// TIA Portal project "ETI C 25" (V15.1) (continued)
   PLC_TO_PC.DATA[324] := ' ';
   PLC_TO_PC.DATA[325] := ' ';
   PLC_TO_PC.DATA[326] := ' ';
   PLC_TO_PC.DATA[327] := ' ';
   PLC_TO_PC.DATA[328] := ' ';
   PLC_TO_PC.DATA[329] := ' ';
   PLC_TO_PC.DATA[330] := ' ';
   PLC_TO_PC.DATA[331] := ' ';
   PLC_TO_PC.DATA[332] := ' ';
   PLC_TO_PC.DATA[333] := ' ';
   PLC_TO_PC.DATA[334] := ' ';
   PLC_TO_PC.DATA[335] := ' ';
   PLC_TO_PC.DATA[336] := ' ';
   PLC_TO_PC.DATA[337] := ' ';
   PLC_TO_PC.DATA[338] := ' ';
   PLC_TO_PC.DATA[339] := ' ';
   PLC_TO_PC.DATA[340] := ' ';
   PLC_TO_PC.DATA[341] := ' ';
   PLC_TO_PC.DATA[342] := ' ';
   PLC_TO_PC.DATA[343] := ' ';
   PLC_TO_PC.DATA[344] := ' ';
   PLC_TO_PC.DATA[345] := ' ';
   PLC_TO_PC.DATA[346] := ' ';
   PLC_TO_PC.DATA[347] := ' ';
   PLC_TO_PC.DATA[348] := ' ';
   PLC_TO_PC.DATA[349] := ' ';
   PLC_TO_PC.DATA[350] := ' ';
   PLC_TO_PC.DATA[351] := ' ';
   PLC_TO_PC.DATA[352] := ' ';
   PLC_TO_PC.DATA[353] := ' ';
   PLC_TO_PC.DATA[354] := ' ';
   PLC_TO_PC.DATA[355] := ' ';
   PLC_TO_PC.DATA[356] := ' ';
   PLC_TO_PC.DATA[357] := ' ';
   PLC_TO_PC.DATA[358] := ' ';
   PLC_TO_PC.DATA[359] := ' ';
   PLC_TO_PC.DATA[360] := ' ';
   PLC_TO_PC.DATA[361] := ' ';
   PLC_TO_PC.DATA[362] := ' ';
   PLC_TO_PC.DATA[363] := ' ';
   PLC_TO_PC.DATA[364] := ' ';
   PLC_TO_PC.DATA[365] := ' ';
   PLC_TO_PC.DATA[366] := ' ';
   PLC_TO_PC.DATA[367] := ' ';
   PLC_TO_PC.DATA[368] := ' ';
   PLC_TO_PC.DATA[369] := ' ';
   PLC_TO_PC.DATA[370] := ' ';
   PLC_TO_PC.DATA[371] := ' ';
   PLC_TO_PC.DATA[372] := ' ';
   PLC_TO_PC.DATA[373] := ' ';
   PLC_TO_PC.DATA[374] := ' ';
   PLC_TO_PC.DATA[375] := ' ';
   PLC_TO_PC.DATA[376] := ' ';
   PLC_TO_PC.DATA[377] := ' ';
   PLC_TO_PC.DATA[378] := ' ';
   PLC_TO_PC.DATA[379] := ' ';
   PLC_TO_PC.DATA[380] := ' ';
   PLC_TO_PC.DATA[381] := ' ';
   PLC_TO_PC.DATA[382] := ' ';
   PLC_TO_PC.DATA[383] := ' ';
   PLC_TO_PC.DATA[384] := ' ';
   PLC_TO_PC.DATA[385] := ' ';
   PLC_TO_PC.DATA[386] := ' ';
   PLC_TO_PC.DATA[387] := ' ';
   PLC_TO_PC.DATA[388] := ' ';
   PLC_TO_PC.DATA[389] := ' ';
   PLC_TO_PC.DATA[390] := ' ';
   PLC_TO_PC.DATA[391] := ' ';
   PLC_TO_PC.DATA[392] := ' ';
   PLC_TO_PC.DATA[393] := ' ';
   PLC_TO_PC.DATA[394] := ' ';
   PLC_TO_PC.DATA[395] := ' ';
   PLC_TO_PC.DATA[396] := ' ';
   PLC_TO_PC.DATA[397] := ' ';
   PLC_TO_PC.DATA[398] := ' ';
   PLC_TO_PC.DATA[399] := ' ';
   PLC_TO_PC.DATA[400] := ' ';
   PLC_TO_PC.DATA[401] := ' ';
   PLC_TO_PC.DATA[402] := ' ';
   PLC_TO_PC.DATA[403] := ' ';
   PLC_TO_PC.DATA[404] := ' ';
   PLC_TO_PC.DATA[405] := ' ';
   PLC_TO_PC.DATA[406] := ' ';
   PLC_TO_PC.DATA[407] := ' ';
   PLC_TO_PC.DATA[408] := ' ';
   PLC_TO_PC.DATA[409] := ' ';
   PLC_TO_PC.DATA[410] := ' ';
   PLC_TO_PC.DATA[411] := ' ';
   PLC_TO_PC.DATA[412] := ' ';
   PLC_TO_PC.DATA[413] := ' ';
   PLC_TO_PC.DATA[414] := ' ';
   PLC_TO_PC.DATA[415] := ' ';
   PLC_TO_PC.DATA[416] := ' ';
   PLC_TO_PC.DATA[417] := ' ';
   PLC_TO_PC.DATA[418] := ' ';
   PLC_TO_PC.DATA[419] := ' ';
   PLC_TO_PC.DATA[420] := ' ';
   PLC_TO_PC.DATA[421] := ' ';
   PLC_TO_PC.DATA[422] := ' ';
   PLC_TO_PC.DATA[423] := ' ';
   PLC_TO_PC.DATA[424] := ' ';
   PLC_TO_PC.DATA[425] := ' ';
   PLC_TO_PC.DATA[426] := ' ';
   PLC_TO_PC.DATA[427] := ' ';
   PLC_TO_PC.DATA[428] := ' ';
   PLC_TO_PC.DATA[429] := ' ';
   PLC_TO_PC.DATA[430] := ' ';
   PLC_TO_PC.DATA[431] := ' ';
   PLC_TO_PC.DATA[432] := ' ';
   PLC_TO_PC.DATA[433] := ' ';
   PLC_TO_PC.DATA[434] := ' ';
   PLC_TO_PC.DATA[435] := ' ';
   PLC_TO_PC.DATA[436] := ' ';
   PLC_TO_PC.DATA[437] := ' ';
   PLC_TO_PC.DATA[438] := ' ';
   PLC_TO_PC.DATA[439] := ' ';
   PLC_TO_PC.DATA[440] := ' ';
   PLC_TO_PC.DATA[441] := ' ';
   PLC_TO_PC.DATA[442] := ' ';
   PLC_TO_PC.DATA[443] := ' ';
   PLC_TO_PC.DATA[444] := ' ';
   PLC_TO_PC.DATA[445] := ' ';
   PLC_TO_PC.DATA[446] := ' ';
   PLC_TO_PC.DATA[447] := ' ';
   PLC_TO_PC.DATA[448] := ' ';
   PLC_TO_PC.DATA[449] := ' ';
   PLC_TO_PC.DATA[450] := ' ';
   PLC_TO_PC.DATA[451] := ' ';
   PLC_TO_PC.DATA[452] := ' ';
   PLC_TO_PC.DATA[453] := ' ';
   PLC_TO_PC.DATA[454] := ' ';
   PLC_TO_PC.DATA[455] := ' ';
   PLC_TO_PC.DATA[456] := ' ';
   PLC_TO_PC.DATA[457] := ' ';
   PLC_TO_PC.DATA[458] := ' ';
   PLC_TO_PC.DATA[459] := ' ';
   PLC_TO_PC.DATA[460] := ' ';
   PLC_TO_PC.DATA[461] := ' ';
   PLC_TO_PC.DATA[462] := ' ';
   PLC_TO_PC.DATA[463] := ' ';
   PLC_TO_PC.DATA[464] := ' ';
   PLC_TO_PC.DATA[465] := ' ';
   PLC_TO_PC.DATA[466] := ' ';
   PLC_TO_PC.DATA[467] := ' ';
   PLC_TO_PC.DATA[468] := ' ';
   PLC_TO_PC.DATA[469] := ' ';
   PLC_TO_PC.DATA[470] := ' ';
   PLC_TO_PC.DATA[471] := ' ';
   PLC_TO_PC.DATA[472] := ' ';
   PLC_TO_PC.DATA[473] := ' ';
   PLC_TO_PC.DATA[474] := ' ';
   PLC_TO_PC.DATA[475] := ' ';
   PLC_TO_PC.DATA[476] := ' ';
   PLC_TO_PC.DATA[477] := ' ';
   PLC_TO_PC.DATA[478] := ' ';
   PLC_TO_PC.DATA[479] := ' ';
   PLC_TO_PC.DATA[480] := ' ';
   PLC_TO_PC.DATA[481] := ' ';
   PLC_TO_PC.DATA[482] := ' ';
   PLC_TO_PC.DATA[483] := ' ';
   PLC_TO_PC.DATA[484] := ' ';
   PLC_TO_PC.DATA[485] := ' ';
   PLC_TO_PC.DATA[486] := ' ';
   PLC_TO_PC.DATA[487] := ' ';
   PLC_TO_PC.DATA[488] := ' ';
   PLC_TO_PC.DATA[489] := ' ';
   PLC_TO_PC.DATA[490] := ' ';
   PLC_TO_PC.DATA[491] := ' ';
   PLC_TO_PC.DATA[492] := ' ';
   PLC_TO_PC.DATA[493] := ' ';
   PLC_TO_PC.DATA[494] := ' ';
   PLC_TO_PC.DATA[495] := ' ';
   PLC_TO_PC.DATA[496] := ' ';
   PLC_TO_PC.DATA[497] := ' ';
   PLC_TO_PC.DATA[498] := ' ';
   PLC_TO_PC.DATA[499] := ' ';
   PLC_TO_PC.DATA[500] := ' ';
   PLC_TO_PC.DATA[501] := ' ';
   PLC_TO_PC.DATA[502] := ' ';
   PLC_TO_PC.DATA[503] := ' ';
   PLC_TO_PC.DATA[504] := ' ';
   PLC_TO_PC.DATA[505] := ' ';
   PLC_TO_PC.DATA[506] := ' ';
   PLC_TO_PC.DATA[507] := ' ';
   PLC_TO_PC.DATA[508] := ' ';
   PLC_TO_PC.DATA[509] := ' ';
   PLC_TO_PC.DATA[510] := ' ';
   PLC_TO_PC.DATA[511] := ' ';
   PLC_TO_PC.DATA[512] := ' ';
   PLC_TO_PC.DATA[513] := ' ';
   PLC_TO_PC.DATA[514] := ' ';
   PLC_TO_PC.DATA[515] := ' ';
   PLC_TO_PC.DATA[516] := ' ';
   PLC_TO_PC.DATA[517] := ' ';
   PLC_TO_PC.DATA[518] := ' ';
   PLC_TO_PC.DATA[519] := ' ';
   PLC_TO_PC.DATA[520] := ' ';
   PLC_TO_PC.DATA[521] := ' ';
   PLC_TO_PC.DATA[522] := ' ';
   PLC_TO_PC.DATA[523] := ' ';
   PLC_TO_PC.DATA[524] := ' ';
   PLC_TO_PC.DATA[525] := ' ';
   PLC_TO_PC.DATA[526] := ' ';
   PLC_TO_PC.DATA[527] := ' ';
   PLC_TO_PC.DATA[528] := ' ';
   PLC_TO_PC.DATA[529] := ' ';
   PLC_TO_PC.DATA[530] := ' ';
   PLC_TO_PC.DATA[531] := ' ';
   PLC_TO_PC.DATA[532] := ' ';
   PLC_TO_PC.DATA[533] := ' ';
   PLC_TO_PC.DATA[534] := ' ';
   PLC_TO_PC.DATA[535] := ' ';
   PLC_TO_PC.DATA[536] := ' ';
   PLC_TO_PC.DATA[537] := ' ';
   PLC_TO_PC.DATA[538] := ' ';
   PLC_TO_PC.DATA[539] := ' ';
   PLC_TO_PC.DATA[540] := ' ';
   PLC_TO_PC.DATA[541] := ' ';
   PLC_TO_PC.DATA[542] := ' ';
   PLC_TO_PC.DATA[543] := ' ';
   PLC_TO_PC.DATA[544] := ' ';
   PLC_TO_PC.DATA[545] := ' ';
   PLC_TO_PC.DATA[546] := ' ';
   PLC_TO_PC.DATA[547] := ' ';
   PLC_TO_PC.DATA[548] := ' ';
   PLC_TO_PC.DATA[549] := ' ';
   PLC_TO_PC.DATA[550] := ' ';
   PLC_TO_PC.DATA[551] := ' ';
   PLC_TO_PC.DATA[552] := ' ';
   PLC_TO_PC.DATA[553] := ' ';
   PLC_TO_PC.DATA[554] := ' ';
   PLC_TO_PC.DATA[555] := ' ';
   PLC_TO_PC.DATA[556] := ' ';
   PLC_TO_PC.DATA[557] := ' ';
   PLC_TO_PC.DATA[558] := ' ';
   PLC_TO_PC.DATA[559] := ' ';
   PLC_TO_PC.DATA[560] := ' ';
   PLC_TO_PC.DATA[561] := ' ';
   PLC_TO_PC.DATA[562] := ' ';
   PLC_TO_PC.DATA[563] := ' ';
   PLC_TO_PC.DATA[564] := ' ';
   PLC_TO_PC.DATA[565] := ' ';
   PLC_TO_PC.DATA[566] := ' ';
   PLC_TO_PC.DATA[567] := ' ';
   PLC_TO_PC.DATA[568] := ' ';
   PLC_TO_PC.DATA[569] := ' ';
   PLC_TO_PC.DATA[570] := ' ';
   PLC_TO_PC.DATA[571] := ' ';
   PLC_TO_PC.DATA[572] := ' ';
   PLC_TO_PC.DATA[573] := ' ';
   PLC_TO_PC.DATA[574] := ' ';
   PLC_TO_PC.DATA[575] := ' ';
   PLC_TO_PC.DATA[576] := ' ';
   PLC_TO_PC.DATA[577] := ' ';
   PLC_TO_PC.DATA[578] := ' ';
   PLC_TO_PC.DATA[579] := ' ';
   PLC_TO_PC.DATA[580] := ' ';
   PLC_TO_PC.DATA[581] := ' ';
   PLC_TO_PC.DATA[582] := ' ';
   PLC_TO_PC.DATA[583] := ' ';
   PLC_TO_PC.DATA[584] := ' ';
   PLC_TO_PC.DATA[585] := ' ';
   PLC_TO_PC.DATA[586] := ' ';
   PLC_TO_PC.DATA[587] := ' ';
   PLC_TO_PC.DATA[588] := ' ';
   PLC_TO_PC.DATA[589] := ' ';
   PLC_TO_PC.DATA[590] := ' ';
   PLC_TO_PC.DATA[591] := ' ';
   PLC_TO_PC.DATA[592] := ' ';
   PLC_TO_PC.DATA[593] := ' ';
   PLC_TO_PC.DATA[594] := ' ';
   PLC_TO_PC.DATA[595] := ' ';
   PLC_TO_PC.DATA[596] := ' ';
   PLC_TO_PC.DATA[597] := ' ';
   PLC_TO_PC.DATA[598] := ' ';
   PLC_TO_PC.DATA[599] := ' ';
   PLC_TO_PC.DATA[600] := ' ';
   PLC_TO_PC.DATA[601] := ' ';
   PLC_TO_PC.DATA[602] := ' ';
   PLC_TO_PC.DATA[603] := ' ';
   PLC_TO_PC.DATA[604] := ' ';
   PLC_TO_PC.DATA[605] := ' ';
   PLC_TO_PC.DATA[606] := ' ';
   PLC_TO_PC.DATA[607] := ' ';
   PLC_TO_PC.DATA[608] := ' ';
   PLC_TO_PC.DATA[609] := ' ';
   PLC_TO_PC.DATA[610] := ' ';
   PLC_TO_PC.DATA[611] := ' ';
   PLC_TO_PC.DATA[612] := ' ';
   PLC_TO_PC.DATA[613] := ' ';
   PLC_TO_PC.DATA[614] := ' ';
   PLC_TO_PC.DATA[615] := ' ';
   PLC_TO_PC.DATA[616] := ' ';
   PLC_TO_PC.DATA[617] := ' ';
   PLC_TO_PC.DATA[618] := ' ';
   PLC_TO_PC.DATA[619] := ' ';
   PLC_TO_PC.DATA[620] := ' ';
   PLC_TO_PC.DATA[621] := ' ';
   PLC_TO_PC.DATA[622] := ' ';
   PLC_TO_PC.DATA[623] := ' ';
   PLC_TO_PC.DATA[624] := ' ';
   PLC_TO_PC.DATA[625] := ' ';
   PLC_TO_PC.DATA[626] := ' ';
   PLC_TO_PC.DATA[627] := ' ';
   PLC_TO_PC.DATA[628] := ' ';
   PLC_TO_PC.DATA[629] := ' ';
   PLC_TO_PC.DATA[630] := ' ';
   PLC_TO_PC.DATA[631] := ' ';
   PLC_TO_PC.DATA[632] := ' ';
   PLC_TO_PC.DATA[633] := ' ';
   PLC_TO_PC.DATA[634] := ' ';
   PLC_TO_PC.DATA[635] := ' ';
   PLC_TO_PC.DATA[636] := ' ';
   PLC_TO_PC.DATA[637] := ' ';
   PLC_TO_PC.DATA[638] := ' ';
   PLC_TO_PC.DATA[639] := ' ';
   PLC_TO_PC.DATA[640] := ' ';
   PLC_TO_PC.DATA[641] := ' ';
   PLC_TO_PC.DATA[642] := ' ';
   PLC_TO_PC.DATA[643] := ' ';
   PLC_TO_PC.DATA[644] := ' ';
   PLC_TO_PC.DATA[645] := ' ';
   PLC_TO_PC.DATA[646] := ' ';
   PLC_TO_PC.DATA[647] := ' ';
   PLC_TO_PC.DATA[648] := ' ';
   PLC_TO_PC.DATA[649] := ' ';
   PLC_TO_PC.DATA[650] := ' ';
   PLC_TO_PC.DATA[651] := ' ';
   PLC_TO_PC.DATA[652] := ' ';
   PLC_TO_PC.DATA[653] := ' ';
   PLC_TO_PC.DATA[654] := ' ';
   PLC_TO_PC.DATA[655] := ' ';
   PLC_TO_PC.DATA[656] := ' ';
   PLC_TO_PC.DATA[657] := ' ';
   PLC_TO_PC.DATA[658] := ' ';
   PLC_TO_PC.DATA[659] := ' ';
   PLC_TO_PC.DATA[660] := ' ';
   PLC_TO_PC.DATA[661] := ' ';
   PLC_TO_PC.DATA[662] := ' ';
   PLC_TO_PC.DATA[663] := ' ';
   PLC_TO_PC.DATA[664] := ' ';
   PLC_TO_PC.DATA[665] := ' ';
   PLC_TO_PC.DATA[666] := ' ';
   PLC_TO_PC.DATA[667] := ' ';
   PLC_TO_PC.DATA[668] := ' ';
   PLC_TO_PC.DATA[669] := ' ';
   PLC_TO_PC.DATA[670] := ' ';
   PLC_TO_PC.DATA[671] := ' ';
   PLC_TO_PC.DATA[672] := ' ';
   PLC_TO_PC.DATA[673] := ' ';
   PLC_TO_PC.DATA[674] := ' ';
   PLC_TO_PC.DATA[675] := ' ';
   PLC_TO_PC.DATA[676] := ' ';
   PLC_TO_PC.DATA[677] := ' ';
   PLC_TO_PC.DATA[678] := ' ';
   PLC_TO_PC.DATA[679] := ' ';
   PLC_TO_PC.DATA[680] := ' ';
   PLC_TO_PC.DATA[681] := ' ';
   PLC_TO_PC.DATA[682] := ' ';
   PLC_TO_PC.DATA[683] := ' ';
   PLC_TO_PC.DATA[684] := ' ';
   PLC_TO_PC.DATA[685] := ' ';
   PLC_TO_PC.DATA[686] := ' ';
   PLC_TO_PC.DATA[687] := ' ';
   PLC_TO_PC.DATA[688] := ' ';
   PLC_TO_PC.DATA[689] := ' ';
   PLC_TO_PC.DATA[690] := ' ';
   PLC_TO_PC.DATA[691] := ' ';
   PLC_TO_PC.DATA[692] := ' ';
   PLC_TO_PC.DATA[693] := ' ';
   PLC_TO_PC.DATA[694] := ' ';
   PLC_TO_PC.DATA[695] := ' ';
   PLC_TO_PC.DATA[696] := ' ';
   PLC_TO_PC.DATA[697] := ' ';
   PLC_TO_PC.DATA[698] := ' ';
   PLC_TO_PC.DATA[699] := ' ';
   PLC_TO_PC.DATA[700] := ' ';
   PLC_TO_PC.DATA[701] := ' ';
   PLC_TO_PC.DATA[702] := ' ';
   PLC_TO_PC.DATA[703] := ' ';
   PLC_TO_PC.DATA[704] := ' ';
   PLC_TO_PC.DATA[705] := ' ';
   PLC_TO_PC.DATA[706] := ' ';
   PLC_TO_PC.DATA[707] := ' ';
   PLC_TO_PC.DATA[708] := ' ';
   PLC_TO_PC.DATA[709] := ' ';
   PLC_TO_PC.DATA[710] := ' ';
   PLC_TO_PC.DATA[711] := ' ';
   PLC_TO_PC.DATA[712] := ' ';
   PLC_TO_PC.DATA[713] := ' ';
   PLC_TO_PC.DATA[714] := ' ';
   PLC_TO_PC.DATA[715] := ' ';
   PLC_TO_PC.DATA[716] := ' ';
   PLC_TO_PC.DATA[717] := ' ';
   PLC_TO_PC.DATA[718] := ' ';
   PLC_TO_PC.DATA[719] := ' ';
   PLC_TO_PC.DATA[720] := ' ';
   PLC_TO_PC.DATA[721] := ' ';
   PLC_TO_PC.DATA[722] := ' ';
   PLC_TO_PC.DATA[723] := ' ';
   PLC_TO_PC.DATA[724] := ' ';
   PLC_TO_PC.DATA[725] := ' ';
   PLC_TO_PC.DATA[726] := ' ';
   PLC_TO_PC.DATA[727] := ' ';
   PLC_TO_PC.DATA[728] := ' ';
   PLC_TO_PC.DATA[729] := ' ';
   PLC_TO_PC.DATA[730] := ' ';
   PLC_TO_PC.DATA[731] := ' ';
   PLC_TO_PC.DATA[732] := ' ';
   PLC_TO_PC.DATA[733] := ' ';
   PLC_TO_PC.DATA[734] := ' ';
   PLC_TO_PC.DATA[735] := ' ';
   PLC_TO_PC.DATA[736] := ' ';
   PLC_TO_PC.DATA[737] := ' ';
   PLC_TO_PC.DATA[738] := ' ';
   PLC_TO_PC.DATA[739] := ' ';
   PLC_TO_PC.DATA[740] := ' ';
   PLC_TO_PC.DATA[741] := ' ';
   PLC_TO_PC.DATA[742] := ' ';
   PLC_TO_PC.DATA[743] := ' ';
   PLC_TO_PC.DATA[744] := ' ';
   PLC_TO_PC.DATA[745] := ' ';
   PLC_TO_PC.DATA[746] := ' ';
   PLC_TO_PC.DATA[747] := ' ';
   PLC_TO_PC.DATA[748] := ' ';
   PLC_TO_PC.DATA[749] := ' ';
   PLC_TO_PC.DATA[750] := ' ';
   PLC_TO_PC.DATA[751] := ' ';
   PLC_TO_PC.DATA[752] := ' ';
   PLC_TO_PC.DATA[753] := ' ';
   PLC_TO_PC.DATA[754] := ' ';
   PLC_TO_PC.DATA[755] := ' ';
   PLC_TO_PC.DATA[756] := ' ';
   PLC_TO_PC.DATA[757] := ' ';
   PLC_TO_PC.DATA[758] := ' ';
   PLC_TO_PC.DATA[759] := ' ';
   PLC_TO_PC.DATA[760] := ' ';
   PLC_TO_PC.DATA[761] := ' ';
   PLC_TO_PC.DATA[762] := ' ';
   PLC_TO_PC.DATA[763] := ' ';
   PLC_TO_PC.DATA[764] := ' ';
   PLC_TO_PC.DATA[765] := ' ';
   PLC_TO_PC.DATA[766] := ' ';
   PLC_TO_PC.DATA[767] := ' ';
   PLC_TO_PC.DATA[768] := ' ';
   PLC_TO_PC.DATA[769] := ' ';
   PLC_TO_PC.DATA[770] := ' ';
   PLC_TO_PC.DATA[771] := ' ';
   PLC_TO_PC.DATA[772] := ' ';
   PLC_TO_PC.DATA[773] := ' ';
   PLC_TO_PC.DATA[774] := ' ';
   PLC_TO_PC.DATA[775] := ' ';
   PLC_TO_PC.DATA[776] := ' ';
   PLC_TO_PC.DATA[777] := ' ';
   PLC_TO_PC.DATA[778] := ' ';
   PLC_TO_PC.DATA[779] := ' ';
   PLC_TO_PC.DATA[780] := ' ';
   PLC_TO_PC.DATA[781] := ' ';
   PLC_TO_PC.DATA[782] := ' ';
   PLC_TO_PC.DATA[783] := ' ';
   PLC_TO_PC.DATA[784] := ' ';
   PLC_TO_PC.DATA[785] := ' ';
   PLC_TO_PC.DATA[786] := ' ';
   PLC_TO_PC.DATA[787] := ' ';
   PLC_TO_PC.DATA[788] := ' ';
   PLC_TO_PC.DATA[789] := ' ';
   PLC_TO_PC.DATA[790] := ' ';
   PLC_TO_PC.DATA[791] := ' ';
   PLC_TO_PC.DATA[792] := ' ';
   PLC_TO_PC.DATA[793] := ' ';
   PLC_TO_PC.DATA[794] := ' ';
   PLC_TO_PC.DATA[795] := ' ';
   PLC_TO_PC.DATA[796] := ' ';
   PLC_TO_PC.DATA[797] := ' ';
   PLC_TO_PC.DATA[798] := ' ';
   PLC_TO_PC.DATA[799] := ' ';
   PLC_TO_PC.DATA[800] := ' ';
   PLC_TO_PC.DATA[801] := ' ';
   PLC_TO_PC.DATA[802] := ' ';
   PLC_TO_PC.DATA[803] := ' ';
   PLC_TO_PC.DATA[804] := ' ';
   PLC_TO_PC.DATA[805] := ' ';
   PLC_TO_PC.DATA[806] := ' ';
   PLC_TO_PC.DATA[807] := ' ';
   PLC_TO_PC.DATA[808] := ' ';
   PLC_TO_PC.DATA[809] := ' ';
   PLC_TO_PC.DATA[810] := ' ';
   PLC_TO_PC.DATA[811] := ' ';
   PLC_TO_PC.DATA[812] := ' ';
   PLC_TO_PC.DATA[813] := ' ';
   PLC_TO_PC.DATA[814] := ' ';
   PLC_TO_PC.DATA[815] := ' ';
   PLC_TO_PC.DATA[816] := ' ';
   PLC_TO_PC.DATA[817] := ' ';
   PLC_TO_PC.DATA[818] := ' ';
   PLC_TO_PC.DATA[819] := ' ';
   PLC_TO_PC.DATA[820] := ' ';
   PLC_TO_PC.DATA[821] := ' ';
   PLC_TO_PC.DATA[822] := ' ';
   PLC_TO_PC.DATA[823] := ' ';
   PLC_TO_PC.DATA[824] := ' ';
   PLC_TO_PC.DATA[825] := ' ';
   PLC_TO_PC.DATA[826] := ' ';
   PLC_TO_PC.DATA[827] := ' ';
   PLC_TO_PC.DATA[828] := ' ';
   PLC_TO_PC.DATA[829] := ' ';
   PLC_TO_PC.DATA[830] := ' ';
   PLC_TO_PC.DATA[831] := ' ';
   PLC_TO_PC.DATA[832] := ' ';
   PLC_TO_PC.DATA[833] := ' ';
   PLC_TO_PC.DATA[834] := ' ';
   PLC_TO_PC.DATA[835] := ' ';
   PLC_TO_PC.DATA[836] := ' ';
   PLC_TO_PC.DATA[837] := ' ';
   PLC_TO_PC.DATA[838] := ' ';
   PLC_TO_PC.DATA[839] := ' ';
   PLC_TO_PC.DATA[840] := ' ';
   PLC_TO_PC.DATA[841] := ' ';
   PLC_TO_PC.DATA[842] := ' ';
   PLC_TO_PC.DATA[843] := ' ';
   PLC_TO_PC.DATA[844] := ' ';
   PLC_TO_PC.DATA[845] := ' ';
   PLC_TO_PC.DATA[846] := ' ';
   PLC_TO_PC.DATA[847] := ' ';
   PLC_TO_PC.DATA[848] := ' ';
   PLC_TO_PC.DATA[849] := ' ';
   PLC_TO_PC.DATA[850] := ' ';
   PLC_TO_PC.DATA[851] := ' ';
   PLC_TO_PC.DATA[852] := ' ';
   PLC_TO_PC.DATA[853] := ' ';
   PLC_TO_PC.DATA[854] := ' ';
   PLC_TO_PC.DATA[855] := ' ';
   PLC_TO_PC.DATA[856] := ' ';
   PLC_TO_PC.DATA[857] := ' ';
   PLC_TO_PC.DATA[858] := ' ';
   PLC_TO_PC.DATA[859] := ' ';
   PLC_TO_PC.DATA[860] := ' ';
   PLC_TO_PC.DATA[861] := ' ';
   PLC_TO_PC.DATA[862] := ' ';
   PLC_TO_PC.DATA[863] := ' ';
   PLC_TO_PC.DATA[864] := ' ';
   PLC_TO_PC.DATA[865] := ' ';
   PLC_TO_PC.DATA[866] := ' ';
   PLC_TO_PC.DATA[867] := ' ';
   PLC_TO_PC.DATA[868] := ' ';
   PLC_TO_PC.DATA[869] := ' ';
   PLC_TO_PC.DATA[870] := ' ';
   PLC_TO_PC.DATA[871] := ' ';
   PLC_TO_PC.DATA[872] := ' ';
   PLC_TO_PC.DATA[873] := ' ';
   PLC_TO_PC.DATA[874] := ' ';
   PLC_TO_PC.DATA[875] := ' ';
   PLC_TO_PC.DATA[876] := ' ';
   PLC_TO_PC.DATA[877] := ' ';
   PLC_TO_PC.DATA[878] := ' ';
   PLC_TO_PC.DATA[879] := ' ';
   PLC_TO_PC.DATA[880] := ' ';
   PLC_TO_PC.DATA[881] := ' ';
   PLC_TO_PC.DATA[882] := ' ';
   PLC_TO_PC.DATA[883] := ' ';
   PLC_TO_PC.DATA[884] := ' ';
   PLC_TO_PC.DATA[885] := ' ';
   PLC_TO_PC.DATA[886] := ' ';
   PLC_TO_PC.DATA[887] := ' ';
   PLC_TO_PC.DATA[888] := ' ';
   PLC_TO_PC.DATA[889] := ' ';
   PLC_TO_PC.DATA[890] := ' ';
   PLC_TO_PC.DATA[891] := ' ';
   PLC_TO_PC.DATA[892] := ' ';
   PLC_TO_PC.DATA[893] := ' ';
   PLC_TO_PC.DATA[894] := ' ';
   PLC_TO_PC.DATA[895] := ' ';
   PLC_TO_PC.DATA[896] := ' ';
   PLC_TO_PC.DATA[897] := ' ';
   PLC_TO_PC.DATA[898] := ' ';
   PLC_TO_PC.DATA[899] := ' ';
   PLC_TO_PC.DATA[900] := ' ';
   PLC_TO_PC.DATA[901] := ' ';
   PLC_TO_PC.DATA[902] := ' ';
   PLC_TO_PC.DATA[903] := ' ';
   PLC_TO_PC.DATA[904] := ' ';
   PLC_TO_PC.DATA[905] := ' ';
   PLC_TO_PC.DATA[906] := ' ';
   PLC_TO_PC.DATA[907] := ' ';
   PLC_TO_PC.DATA[908] := ' ';
   PLC_TO_PC.DATA[909] := ' ';
   PLC_TO_PC.DATA[910] := ' ';
   PLC_TO_PC.DATA[911] := ' ';
   PLC_TO_PC.DATA[912] := ' ';
   PLC_TO_PC.DATA[913] := ' ';
   PLC_TO_PC.DATA[914] := ' ';
   PLC_TO_PC.DATA[915] := ' ';
   PLC_TO_PC.DATA[916] := ' ';
   PLC_TO_PC.DATA[917] := ' ';
   PLC_TO_PC.DATA[918] := ' ';
   PLC_TO_PC.DATA[919] := ' ';
   PLC_TO_PC.DATA[920] := ' ';
   PLC_TO_PC.DATA[921] := ' ';
   PLC_TO_PC.DATA[922] := ' ';
   PLC_TO_PC.DATA[923] := ' ';
   PLC_TO_PC.DATA[924] := ' ';
   PLC_TO_PC.DATA[925] := ' ';
   PLC_TO_PC.DATA[926] := ' ';
   PLC_TO_PC.DATA[927] := ' ';
   PLC_TO_PC.DATA[928] := ' ';
   PLC_TO_PC.DATA[929] := ' ';
   PLC_TO_PC.DATA[930] := ' ';
   PLC_TO_PC.DATA[931] := ' ';
   PLC_TO_PC.DATA[932] := ' ';
   PLC_TO_PC.DATA[933] := ' ';
   PLC_TO_PC.DATA[934] := ' ';
   PLC_TO_PC.DATA[935] := ' ';
   PLC_TO_PC.DATA[936] := ' ';
   PLC_TO_PC.DATA[937] := ' ';
   PLC_TO_PC.DATA[938] := ' ';
   PLC_TO_PC.DATA[939] := ' ';
   PLC_TO_PC.DATA[940] := ' ';
   PLC_TO_PC.DATA[941] := ' ';
   PLC_TO_PC.DATA[942] := ' ';
   PLC_TO_PC.DATA[943] := ' ';
   PLC_TO_PC.DATA[944] := ' ';
   PLC_TO_PC.DATA[945] := ' ';
   PLC_TO_PC.DATA[946] := ' ';
   PLC_TO_PC.DATA[947] := ' ';
   PLC_TO_PC.DATA[948] := ' ';
   PLC_TO_PC.DATA[949] := ' ';
   PLC_TO_PC.DATA[950] := ' ';
   PLC_TO_PC.DATA[951] := ' ';
   PLC_TO_PC.DATA[952] := ' ';
   PLC_TO_PC.DATA[953] := ' ';
   PLC_TO_PC.DATA[954] := ' ';
   PLC_TO_PC.DATA[955] := ' ';
   PLC_TO_PC.DATA[956] := ' ';
   PLC_TO_PC.DATA[957] := ' ';
   PLC_TO_PC.DATA[958] := ' ';
   PLC_TO_PC.DATA[959] := ' ';
   PLC_TO_PC.DATA[960] := ' ';
   PLC_TO_PC.DATA[961] := ' ';
   PLC_TO_PC.DATA[962] := ' ';
   PLC_TO_PC.DATA[963] := ' ';
   PLC_TO_PC.DATA[964] := ' ';
   PLC_TO_PC.DATA[965] := ' ';
   PLC_TO_PC.DATA[966] := ' ';
   PLC_TO_PC.DATA[967] := ' ';
   PLC_TO_PC.DATA[968] := ' ';
   PLC_TO_PC.DATA[969] := ' ';
   PLC_TO_PC.DATA[970] := ' ';
   PLC_TO_PC.DATA[971] := ' ';
   PLC_TO_PC.DATA[972] := ' ';
   PLC_TO_PC.DATA[973] := ' ';
   PLC_TO_PC.DATA[974] := ' ';
   PLC_TO_PC.DATA[975] := ' ';
   PLC_TO_PC.DATA[976] := ' ';
   PLC_TO_PC.DATA[977] := ' ';
   PLC_TO_PC.DATA[978] := ' ';
   PLC_TO_PC.DATA[979] := ' ';
   PLC_TO_PC.DATA[980] := ' ';
   PLC_TO_PC.DATA[981] := ' ';
   PLC_TO_PC.DATA[982] := ' ';
   PLC_TO_PC.DATA[983] := ' ';
   PLC_TO_PC.DATA[984] := ' ';
   PLC_TO_PC.DATA[985] := ' ';
   PLC_TO_PC.DATA[986] := ' ';
   PLC_TO_PC.DATA[987] := ' ';
   PLC_TO_PC.DATA[988] := ' ';
   PLC_TO_PC.DATA[989] := ' ';
   PLC_TO_PC.DATA[990] := ' ';
   PLC_TO_PC.DATA[991] := ' ';
   PLC_TO_PC.DATA[992] := ' ';
   PLC_TO_PC.DATA[993] := ' ';
   PLC_TO_PC.DATA[994] := ' ';
   PLC_TO_PC.DATA[995] := ' ';
   PLC_TO_PC.DATA[996] := ' ';
   PLC_TO_PC.DATA[997] := ' ';
   PLC_TO_PC.DATA[998] := ' ';
   PLC_TO_PC.DATA[999] := ' ';
   PLC_TO_PC.DATA[1000] := ' ';
   PLC_TO_PC.DATA[1001] := ' ';
   PLC_TO_PC.DATA[1002] := ' ';
   PLC_TO_PC.DATA[1003] := ' ';
   PLC_TO_PC.DATA[1004] := ' ';
   PLC_TO_PC.DATA[1005] := ' ';
   PLC_TO_PC.DATA[1006] := ' ';
   PLC_TO_PC.DATA[1007] := ' ';
   PLC_TO_PC.DATA[1008] := ' ';
   PLC_TO_PC.DATA[1009] := ' ';
   PLC_TO_PC.DATA[1010] := ' ';
   PLC_TO_PC.DATA[1011] := ' ';
   PLC_TO_PC.DATA[1012] := ' ';
   PLC_TO_PC.DATA[1013] := ' ';
   PLC_TO_PC.DATA[1014] := ' ';
   PLC_TO_PC.DATA[1015] := ' ';
   PLC_TO_PC.DATA[1016] := ' ';
   PLC_TO_PC.DATA[1017] := ' ';
   PLC_TO_PC.DATA[1018] := ' ';
   PLC_TO_PC.DATA[1019] := ' ';
   PLC_TO_PC.DATA[1020] := ' ';
   PLC_TO_PC.DATA[1021] := ' ';
   PLC_TO_PC.DATA[1022] := ' ';
   PLC_TO_PC.DATA[1023] := ' ';
END_DATA_BLOCK

DATA_BLOCK "FB_Lin_fun_DB_FB_SDAT"   // DB18
{ S7_Optimized_Access := 'TRUE' }
VERSION : 0.1
// stored: InstanceOfName FB_Lin_fun
"FB_Lin_fun"
BEGIN
END_DATA_BLOCK

DATA_BLOCK "DB_KEYENCE"   // DB19
{ S7_Optimized_Access := 'TRUE' }
VERSION : 0.1
   VAR RETAIN
      Elektroda : Struct
         ZeljenaPozicija : Struct
            POZ1_elektrodaGor : UInt := 58700;   // ELektrodaOdmik
            POZ2_elektrodaVmes : UInt := 0;   // Elektroda odmaknjena
            POZ3_elektrodaStisnjena : UInt := 37100;   // ElektrodaStisnjena
            POZ4_elektrodaZavarjeno : UInt := 0;   // ElektrodaVPozicijiZavarjeno
         END_STRUCT;
         HISTEREZA : UInt := 600;
         TOLERANCA : Array[1..4] of Int;
      END_STRUCT;
      Kroznik : Struct
         ZeljenaPozicija : Struct
            POZ1_KonusNazaj : UInt := 60000;   // KonusSproscen
            POZ2_KonusNaprej : UInt := 56840;   // KonusZaprt
         END_STRUCT;
      END_STRUCT;
      HSTEREZA : UInt := 400;
      TOLERANCA : Array[1..4] of Int;
   END_VAR
BEGIN
END_DATA_BLOCK

DATA_BLOCK "FB_KEYENCE_GT2_ODMIKVARJENJA"   // DB20
{ S7_Optimized_Access := 'TRUE' }
VERSION : 0.1
// stored: InstanceOfName FB_KEYENCE_GT2
"FB_KEYENCE_GT2"
BEGIN
END_DATA_BLOCK

DATA_BLOCK "FB_KEYENCE_GT2_odmikKonusaKroznika"   // DB21
{ S7_Optimized_Access := 'TRUE' }
VERSION : 0.1
// stored: InstanceOfName FB_KEYENCE_GT2
"FB_KEYENCE_GT2"
BEGIN
END_DATA_BLOCK

DATA_BLOCK "FB_AKD_VrtenjeKroznika"   // DB22
{ S7_Optimized_Access := 'TRUE' }
VERSION : 0.1
// stored: InstanceOfName FB_AKD
"FB_AKD"
BEGIN
END_DATA_BLOCK

DATA_BLOCK "FB_AKD_VrtenjeELektrode"   // DB23
{ S7_Optimized_Access := 'TRUE' }
VERSION : 0.1
// stored: InstanceOfName FB_AKD
"FB_AKD"
BEGIN
END_DATA_BLOCK

DATA_BLOCK "FB_AKD_DB_elektroda"   // DB24
{ S7_Optimized_Access := 'TRUE' }
VERSION : 0.1
// stored: InstanceOfName FB_AKD
"FB_AKD"
BEGIN
END_DATA_BLOCK

DATA_BLOCK "FB_AKD_DB"   // DB25
{ S7_Optimized_Access := 'TRUE' }
VERSION : 0.1
// stored: InstanceOfName FB_AKD
"FB_AKD"
BEGIN
END_DATA_BLOCK

DATA_BLOCK "FB_AKD_DB_RezanjePodajanje"   // DB28
{ S7_Optimized_Access := 'TRUE' }
VERSION : 0.1
// stored: InstanceOfName FB_AKD
"FB_AKD"
BEGIN
END_DATA_BLOCK

DATA_BLOCK "DB_PODATKI"   // DB29
{ S7_Optimized_Access := 'TRUE' }
VERSION : 0.1
   VAR RETAIN
      KROZNA_MIZA : Struct
         IzdelekPrisoten : Byte;
         IzdelekZavarjen : Byte;
         IzdelekKameraOk : Byte;
         merkerjiprisotnost : Array[0..1] of Bool;
         merkerjivarjenje : Array[0..10] of Bool;
         merkerjiIzmeta : Array[0..10] of Bool;
         IzdelekPrisotenArray : Array[0..7] of Bool;
         StatusIzdelkaVarjenje : Array[0..7] of Byte;
         StatusIzdelkaKamera : Array[0..7] of Byte;
         MerkerjiKoraka : Array[0..100] of Bool;
      END_STRUCT;
      GeaphName : String := 'FB_GL_PROGRAM';
      HMI_ALARM : WString;
   END_VAR
   VAR
      StartupBit : Bool;
      StartupbitMerker : Bool;
   END_VAR
   VAR RETAIN
      Merkerji_OdvijanjeTraku_Ciscenje : Array[0..9] of Bool;
   END_VAR
BEGIN
END_DATA_BLOCK

DATA_BLOCK "FB_IZMETKOMADA_DB"   // DB30
{ S7_Optimized_Access := 'TRUE' }
VERSION : 0.1
// stored: InstanceOfName FB_IZMETKOMADA
"FB_IZMETKOMADA"
BEGIN
END_DATA_BLOCK

DATA_BLOCK "DB_VARJENJE"   // DB35
{ S7_Optimized_Access := 'TRUE' }
VERSION : 0.1
   VAR RETAIN
      PODATKI : Struct
         input : Struct
            ZajtevaZaVarjenje : Bool := FALSE;
            IzbiraPrograma : Byte := 16#05;
            VarilniTokOn : Bool := TRUE;
            SpotSelectionOn : Bool := TRUE;
         END_STRUCT;
         TON_timers : Array[0..1] of TON_TIME;
         TP_timers : Array[0..1] of TP_TIME;
         VarjenjeON : Bool := TRUE;
      END_STRUCT;
      merkerji : Array[0..1] of Bool;
   END_VAR
BEGIN
   PODATKI.TON_timers[0].ST := T#0MS;
   PODATKI.TON_timers[0].PT := T#0MS;
   PODATKI.TON_timers[0].RU := FALSE;
   PODATKI.TON_timers[0].IN := FALSE;
   PODATKI.TON_timers[1].ST := T#0MS;
   PODATKI.TON_timers[1].PT := T#0MS;
   PODATKI.TON_timers[1].RU := FALSE;
   PODATKI.TON_timers[1].IN := FALSE;
   PODATKI.TP_timers[0].ST := T#0MS;
   PODATKI.TP_timers[0].PT := T#0MS;
   PODATKI.TP_timers[0].RU := FALSE;
   PODATKI.TP_timers[0].IN := FALSE;
   PODATKI.TP_timers[1].ST := T#0MS;
   PODATKI.TP_timers[1].PT := T#0MS;
   PODATKI.TP_timers[1].RU := FALSE;
   PODATKI.TP_timers[1].IN := FALSE;
   merkerji[0] := FALSE;
   merkerji[1] := FALSE;
   // PODATKI.TON_timers[0] : TImer pulz varjenja
END_DATA_BLOCK

DATA_BLOCK "FB_Alarms_DB"   // DB37
{ S7_Optimized_Access := 'TRUE' }
AUTHOR : Andrej
VERSION : 0.1
// stored: InstanceOfName FB_Alarms
"FB_Alarms"
BEGIN
END_DATA_BLOCK

DATA_BLOCK "GRAPH_HMI"   // DB38
{ S7_Optimized_Access := 'FALSE' }
VERSION : 0.1
   VAR
      HMINAME : Array[0..254] of String;
   END_VAR
BEGIN
END_DATA_BLOCK

DATA_BLOCK "MERJERJI"   // DB39
{ S7_Optimized_Access := 'TRUE' }
VERSION : 0.1
   VAR RETAIN
      merjer : Array[0..250] of Bool;
   END_VAR
BEGIN
END_DATA_BLOCK

DATA_BLOCK "FB_VstavljanjeIzdelkaVMizo_DB"   // DB40
{ S7_Optimized_Access := 'TRUE' }
VERSION : 0.1
// stored: InstanceOfName FB_VstavljanjeIzdelkaVMizo
"FB_VstavljanjeIzdelkaVMizo"
BEGIN
END_DATA_BLOCK

DATA_BLOCK "FB_Alarms_DB_1"   // DB42
{ S7_Optimized_Access := 'TRUE' }
AUTHOR : Andrej
VERSION : 0.1
// stored: InstanceOfName FB_Alarms
"FB_Alarms"
BEGIN
END_DATA_BLOCK

DATA_BLOCK "FB_IOL_BANNER_DB"   // DB46
{ S7_Optimized_Access := 'TRUE' }
VERSION : 0.1
// stored: InstanceOfName FB_IOL_BANNER
"FB_IOL_BANNER"
BEGIN
END_DATA_BLOCK

DATA_BLOCK "DB_IOL_BANNER"   // DB47
{ S7_Optimized_Access := 'TRUE' }
VERSION : 0.1
   VAR RETAIN
      PODATKI : Struct
         Color1 : Byte;
         ColorFlashRange : Byte;
         Color2 : Byte;
         AdiableMode : Byte;
         CV : Bool;
         AnimationType : Byte;
         Color1Intensity : Byte;
         Color2Intensity : Byte;
      END_STRUCT;
   END_VAR
BEGIN
END_DATA_BLOCK

DATA_BLOCK "DB_STEVCI"   // DB56
{ S7_Optimized_Access := 'TRUE' }
VERSION : 0.1
   VAR RETAIN
      "STEVCI VARJENJE" : Struct
         ZavarjenoOK : UInt;
         ZavarjenoNOK : UInt;
         SKUPAJOK : UInt;
         SKUPAJNOK : UInt;
         SKUPAJ : UInt;
      END_STRUCT;
      "STEVCI KAMERA" : Struct
         KameraOK : UInt;
         KameraNOK : UInt;
         SKUPAJOK : UInt;
         SKUPAJNOK : UInt;
         SKUPAJ : UInt;
      END_STRUCT;
      STEVEC_SKATEL : Struct
         SKATLA1 : UInt;
         SKATLA2 : UInt;
         SKATLA_SLABI : UInt;
      END_STRUCT;
      STEVCI_ZELENAPOLNA_SKATLA : Struct
         SKATLA1 : UInt := 1300;
         SKATLA2 : UInt := 1300;
         skatla1polna : Bool;
         skatla2polna : Bool;
         skatlaslabi : UInt := 20;
         merkerji : Array[0..1] of Bool;
      END_STRUCT;
      STEVEC_PREKLOPOV : UInt;
      bacSTEVEC_PREKLOPOV : UInt;
      nCounterOdvijanjeTrakuCiscenje : DInt;
   END_VAR
BEGIN
END_DATA_BLOCK

DATA_BLOCK "FB_TekociTrak_DB"   // DB59
{ S7_Optimized_Access := 'TRUE' }
VERSION : 0.1
// stored: InstanceOfName FB_TekociTrak
"FB_TekociTrak"
BEGIN
END_DATA_BLOCK

DATA_BLOCK "FB_CYCLETIME"   // DB62
{ S7_Optimized_Access := 'TRUE' }
VERSION : 0.1
// stored: InstanceOfName FB_TIMERS
"FB_TIMERS"
BEGIN
END_DATA_BLOCK

DATA_BLOCK "Block_1_DB"   // DB65
{ S7_Optimized_Access := 'TRUE' }
VERSION : 0.1
// stored: InstanceOfName Block_1
"Block_1"
BEGIN
END_DATA_BLOCK

DATA_BLOCK "FB_LocalTime_DB"   // DB66
{ S7_Optimized_Access := 'TRUE' }
VERSION : 0.1
// stored: InstanceOfName FB_LocalTime
"FB_LocalTime"
BEGIN
END_DATA_BLOCK

DATA_BLOCK "FB_KAMERA_TRIG_DB"   // DB67
{ S7_Optimized_Access := 'TRUE' }
VERSION : 0.1
// stored: InstanceOfName FB_KAMERA_TRIG
"FB_KAMERA_TRIG"
BEGIN
END_DATA_BLOCK

// folder: System blocks/Program resources

DATA_BLOCK "IEC_Timer_0_DB"   // DB7
{ S7_Optimized_Access := 'TRUE' }
AUTHOR : Simatic
FAMILY : IEC
NAME : IEC_TMR
VERSION : 1.0
// stored: InstanceOfName IEC_TIMER
"IEC_TIMER"
BEGIN
END_DATA_BLOCK

DATA_BLOCK "PLC_1_Connection_DB"   // DB27
{ S7_Optimized_Access := 'TRUE' }
AUTHOR : SIMATIC
FAMILY : MC7Plus
NAME : TC_IP_v4
VERSION : 1.0
// stored: InstanceOfName TCON_IP_v4
"TCON_IP_v4"
BEGIN
   ID := 1;
   InterfaceId := 64;
   LocalPort := 4999;
   RemotePort := 5000;
   ActiveEstablished := true;
   RemoteAddress.ADDR[1] := 192;
   RemoteAddress.ADDR[2] := 168;
   RemoteAddress.ADDR[4] := 200;
END_DATA_BLOCK

DATA_BLOCK "TON_MOTOR"   // DB31
{ S7_Optimized_Access := 'TRUE' }
AUTHOR : Simatic
FAMILY : IEC
NAME : IEC_TMR
VERSION : 1.0
// stored: InstanceOfName IEC_TIMER
"IEC_TIMER"
BEGIN
END_DATA_BLOCK

DATA_BLOCK "TImerPodajanja"   // DB32
{ S7_Optimized_Access := 'TRUE' }
AUTHOR : Simatic
FAMILY : IEC
NAME : IEC_TMR
VERSION : 1.0
// stored: InstanceOfName IEC_TIMER
"IEC_TIMER"
BEGIN
END_DATA_BLOCK

DATA_BLOCK "IEC_Timer_0_DB_1"   // DB33
{ S7_Optimized_Access := 'TRUE' }
AUTHOR : Simatic
FAMILY : IEC
NAME : IEC_TMR
VERSION : 1.0
// stored: InstanceOfName IEC_TIMER
"IEC_TIMER"
BEGIN
END_DATA_BLOCK

DATA_BLOCK "TON_REZANJEPODAJANJE"   // DB34
{ S7_Optimized_Access := 'TRUE' }
AUTHOR : Simatic
FAMILY : IEC
NAME : IEC_TMR
VERSION : 1.0
// stored: InstanceOfName IEC_TIMER
"IEC_TIMER"
BEGIN
END_DATA_BLOCK

DATA_BLOCK "IEC_Timer_0_DB_2"   // DB36
{ S7_Optimized_Access := 'TRUE' }
AUTHOR : Simatic
FAMILY : IEC
NAME : IEC_TMR
VERSION : 1.0
// stored: InstanceOfName IEC_TIMER
"IEC_TIMER"
BEGIN
END_DATA_BLOCK

DATA_BLOCK "IEC_Timer_0_DB_3"   // DB41
{ S7_Optimized_Access := 'TRUE' }
AUTHOR : Simatic
FAMILY : IEC
NAME : IEC_TMR
VERSION : 1.0
// stored: InstanceOfName IEC_TIMER
"IEC_TIMER"
BEGIN
END_DATA_BLOCK

DATA_BLOCK "TON_UDP_STARTUP"   // DB45
{ S7_Optimized_Access := 'TRUE' }
AUTHOR : Simatic
FAMILY : IEC
NAME : IEC_TMR
VERSION : 1.0
// stored: InstanceOfName IEC_TIMER
"IEC_TIMER"
BEGIN
END_DATA_BLOCK

DATA_BLOCK "STEVECKOSOV_PO_KONCU_TRAKU"   // DB48
{ S7_Optimized_Access := 'TRUE' }
AUTHOR : Simatic
FAMILY : IEC
NAME : CNTR
VERSION : 1.0
// stored: InstanceOfName IEC_COUNTER
"IEC_COUNTER"
BEGIN
END_DATA_BLOCK

DATA_BLOCK "IEC_Timer_0_DB_5"   // DB49
{ S7_Optimized_Access := 'TRUE' }
AUTHOR : Simatic
FAMILY : IEC
NAME : IEC_TMR
VERSION : 1.0
// stored: InstanceOfName IEC_TIMER
"IEC_TIMER"
BEGIN
END_DATA_BLOCK

DATA_BLOCK "IEC_Timer_0_DB_4"   // DB50
{ S7_Optimized_Access := 'TRUE' }
AUTHOR : Simatic
FAMILY : IEC
NAME : IEC_TMR
VERSION : 1.0
// stored: InstanceOfName IEC_TIMER
"IEC_TIMER"
BEGIN
END_DATA_BLOCK

DATA_BLOCK "IEC_Timer_0_DB_6"   // DB51
{ S7_Optimized_Access := 'TRUE' }
AUTHOR : Simatic
FAMILY : IEC
NAME : IEC_TMR
VERSION : 1.0
// stored: InstanceOfName IEC_TIMER
"IEC_TIMER"
BEGIN
END_DATA_BLOCK

DATA_BLOCK "IEC_Timer_0_DB_7"   // DB52
{ S7_Optimized_Access := 'TRUE' }
AUTHOR : Simatic
FAMILY : IEC
NAME : IEC_TMR
VERSION : 1.0
// stored: InstanceOfName IEC_TIMER
"IEC_TIMER"
BEGIN
END_DATA_BLOCK

DATA_BLOCK "IEC_Timer_0_DB_8"   // DB53
{ S7_Optimized_Access := 'TRUE' }
AUTHOR : Simatic
FAMILY : IEC
NAME : IEC_TMR
VERSION : 1.0
// stored: InstanceOfName IEC_TIMER
"IEC_TIMER"
BEGIN
END_DATA_BLOCK

DATA_BLOCK "IEC_Timer_0_DB_9"   // DB54
{ S7_Optimized_Access := 'TRUE' }
AUTHOR : Simatic
FAMILY : IEC
NAME : IEC_TMR
VERSION : 1.0
// stored: InstanceOfName IEC_TIMER
"IEC_TIMER"
BEGIN
END_DATA_BLOCK

DATA_BLOCK "IEC_Timer_0_DB_10"   // DB55
{ S7_Optimized_Access := 'TRUE' }
AUTHOR : Simatic
FAMILY : IEC
NAME : IEC_TMR
VERSION : 1.0
// stored: InstanceOfName IEC_TIMER
"IEC_TIMER"
BEGIN
END_DATA_BLOCK

DATA_BLOCK "IEC_Timer_0_DB_11"   // DB57
{ S7_Optimized_Access := 'TRUE' }
AUTHOR : Simatic
FAMILY : IEC
NAME : IEC_TMR
VERSION : 1.0
// stored: InstanceOfName IEC_TIMER
"IEC_TIMER"
BEGIN
END_DATA_BLOCK

DATA_BLOCK "IEC_Counter_0_DB"   // DB58
{ S7_Optimized_Access := 'TRUE' }
AUTHOR : Simatic
FAMILY : IEC
NAME : UCNTR
VERSION : 1.2
// stored: InstanceOfName IEC_UCOUNTER
"IEC_UCOUNTER"
BEGIN
END_DATA_BLOCK

DATA_BLOCK "IEC_Timer_0_DB_12"   // DB60
{ S7_Optimized_Access := 'TRUE' }
AUTHOR : Simatic
FAMILY : IEC
NAME : IEC_TMR
VERSION : 1.0
// stored: InstanceOfName IEC_TIMER
"IEC_TIMER"
BEGIN
END_DATA_BLOCK

DATA_BLOCK "IEC_Timer_0_DB_13"   // DB61
{ S7_Optimized_Access := 'TRUE' }
AUTHOR : Simatic
FAMILY : IEC
NAME : IEC_TMR
VERSION : 1.0
// stored: InstanceOfName IEC_TIMER
"IEC_TIMER"
BEGIN
END_DATA_BLOCK

DATA_BLOCK "IEC_Counter_0_DB_1"   // DB64
{ S7_Optimized_Access := 'TRUE' }
AUTHOR : Simatic
FAMILY : IEC
NAME : CNTR
VERSION : 1.0
// stored: InstanceOfName IEC_COUNTER
"IEC_COUNTER"
BEGIN
END_DATA_BLOCK

DATA_BLOCK "IEC_Timer_0_DB_15"   // DB68
{ S7_Optimized_Access := 'TRUE' }
AUTHOR : Simatic
FAMILY : IEC
NAME : IEC_TMR
VERSION : 1.0
// stored: InstanceOfName IEC_TIMER
"IEC_TIMER"
BEGIN
END_DATA_BLOCK

// folder: (top level)

FUNCTION_BLOCK "FB_IOL_SDAT"   // FB1, LAD
{ S7_Optimized_Access := 'TRUE' }
VERSION : 0.1
// VHOD : DWord naslov IOL linka
// 
// Blok pretvori vhodne podatke v izhodno vrednost in posatavi bite za končne položaje (bBDC1- bBDC4)
   VAR_INPUT
      w_inAddr : Word;   // VALUE| VALUE|VALUE|BDC1-4
      iPoz1 : Real;
      iPoz2 : Real;
      iPoz3 : Real;
      iPoz4 : Real;
      Histereza : Real := 0.1;
   END_VAR
   VAR_OUTPUT
      out : Real;   // Rezultat int
      bBDC1 : Bool;   // Končni položaj 1
      bBDC2 : Bool;   // Končni položaj 2
      bBDC3 : Bool;   // Končni položaj 3
      bBDC4 : Bool;   // Končni položaj 4
      oPoz1Dosezena : Bool;
      oPoz2Dosezena : Bool;
      oPoz3Dosezena : Bool;
      oPoz4Dosezena : Bool;
   END_VAR
   VAR RETAIN
      w_statRor : Word;
      W_ST : Word;
   END_VAR
   VAR
      B0 : Byte;
      B1 : Byte;
      FB_Lin_fun_Instance : "FB_Lin_fun";
   END_VAR
   VAR_TEMP
      temp1 : Real;
   END_VAR
BEGIN

REGION Network 2 (SCL)
   #B0 := #w_inAddr.%B0;
   #B1 := #w_inAddr.%B1;

   //#W_ST := SWAP(#w_inAddr);
   //Rotacija za 4 bite v desno |PODATKI|PODATKI| PODATKI|BDC1-BDC4|
   //Rezultat b0-b12 predstavlja rezultat
   #w_statRor := SHR(IN := #w_inAddr, N := 4);

   //maskiramo samo prvih 12 bitov 16#0FFF; 
   #temp1 :=UINT_TO_REAL(( #w_statRor AND 2#0000_1111_1111_1111));
   //resolucija 0.05mm

   #FB_Lin_fun_Instance(I_PIW_real:=#temp1,
                        I_x2:=1679.0,
                        I_x1:=0.0,
                        I_y2:=80.0,
                        I_y1:=0.0);


   #out := #FB_Lin_fun_Instance.Q_izhod;

   //zadnje 4 bite uproabimo za BDC indikacijo
   #bBDC1 := #w_statRor.%X12;
   #bBDC1 := #w_statRor.%X13;
   #bBDC1 := #w_statRor.%X14;
   #bBDC1 := #w_statRor.%X15;
END_REGION

REGION Network 3 (SCL)
   //pozicija dosezena
   //
   IF (#iPoz1 - #Histereza) < #out AND #out < (#iPoz1 + #Histereza) AND #iPoz1 <> 0  THEN
       #oPoz1Dosezena := true;
   ELSE
       #oPoz1Dosezena := false;
   END_IF;

   IF (#iPoz2 - #Histereza) < #out AND #out < (#iPoz2 + #Histereza) AND #iPoz1 <> 0 THEN
       #oPoz2Dosezena := true;
   ELSE
       #oPoz2Dosezena := false;
   END_IF;
END_REGION
END_FUNCTION_BLOCK

FUNCTION_BLOCK "FB_MVK1"   // FB2, LAD
{ S7_Optimized_Access := 'TRUE' }
VERSION : 0.1
   VAR_INPUT
      myWORD : Word;
   END_VAR
   VAR
      stat_myWord : Word;
   END_VAR
   VAR RETAIN
      Senzorji : "UDT_MVK1";
   END_VAR
BEGIN

REGION Network 2
   // xc
END_REGION

REGION Network 3 (SCL)
   #stat_myWord := ROR(IN:=#myWORD, N:=8);

   #Senzorji."1Y1".B1 := #stat_myWord.%X0;
   #Senzorji."1Y1".B2 := #stat_myWord.%X1;
END_REGION
END_FUNCTION_BLOCK

FUNCTION_BLOCK "FB_IOL_IFM_SV"   // FB3, SCL
{ S7_Optimized_Access := 'TRUE' }
VERSION : 0.1
   VAR_INPUT
      d_slaveAddr : DWord;   // Nalov IOL slave naprave - 4 byte
      iminZeljeniPretok : UInt;
      iMaxTeperautra : Real;
   END_VAR
   VAR_OUTPUT
      BDC1 : Bool;
      BDC2 : Bool;
      uPretok : UInt;
      fTemperatura : Real;
      oPretokOK : Bool;
      oTempOK : Bool;
   END_VAR
   VAR RETAIN
      d_slaveValue : DWord;   // Vrednost na IOL naslovu
      B_slaveByte : Array[0..3] of Word;
   END_VAR
   VAR
      stat_iTemperatura : Int;
      stat_uPretok : UInt;
   END_VAR
BEGIN
   (*
   PROGRAMSKI BLOK ZA IOL LINK
   SLAVE : IFM - SV serija - merilniki pretoka

   IN : WORD
   OUT : BDC1
       : BDC2
       : Temperatura
       : Pretok
   *)

   //prepis v statični del pomnilnika
   #d_slaveValue := #d_slaveAddr;


   //menjava High and Low byta - IOL -> profinet big Endian
   #B_slaveByte[0] := #d_slaveValue.%B0;
   #B_slaveByte[1] := #d_slaveValue.%B1;
   #B_slaveByte[2] := #d_slaveValue.%B2;
   #B_slaveByte[3] := #d_slaveValue.%B3;

   //0 bit - BDC1
   #BDC1 := #B_slaveByte[0].%X0;
   //1 bit - BDC2
   #BDC2 := #B_slaveByte[0].%X1;

   //Merjenje temperature
   #stat_iTemperatura := SHL(IN:=#B_slaveByte[1],N:=8)+ #B_slaveByte[0];
   //zmakni meritev za 2 bita
   #stat_iTemperatura := SHR(IN := #stat_iTemperatura, N := 2);
   //pretvori v float vrednost
   #fTemperatura := #stat_iTemperatura / 10.0;


   //#B_slaveByte[]
   //#u_Pretok := 16#0000_0000 + (SHL(IN:=
   #stat_uPretok := SHL(IN := #B_slaveByte[3], N := 8) + #B_slaveByte[2];
   #uPretok := #stat_uPretok;

   IF #uPretok>#iminZeljeniPretok THEN
       #oPretokOK := true;
   ELSE
       #oPretokOK := false;
   END_IF;

   IF #iMaxTeperautra > #iminZeljeniPretok THEN
       #oTempOK := true;
   ELSE
       #oTempOK := false;
   END_IF;
END_FUNCTION_BLOCK

FUNCTION_BLOCK "FB_FESTO_VPPM"   // FB4, SCL
{ S7_Optimized_Access := 'TRUE' }
VERSION : 0.1
   VAR_INPUT
      addrTrenutniPritisk : Word;
   END_VAR
   VAR_OUTPUT
      TrenutniPritisk : Real;
      SetPoint : UInt;
      PritiskDosezen : Bool;
   END_VAR
   VAR RETAIN
      statZeleniPritisk : Int;
      setstatZeljeniPritisk : Real;
   END_VAR
BEGIN
   #TrenutniPritisk := #addrTrenutniPritisk / 1000.0;
   #statZeleniPritisk :=  #setstatZeljeniPritisk * 1000;
   #SetPoint := UINT_TO_WORD(IN:=#statZeleniPritisk);
   //#SetPoint := ROR(IN := #SetPoint,N:=8);
   //

   IF #SetPoint = #TrenutniPritisk THEN
       #PritiskDosezen := true;
   ELSE
       #PritiskDosezen := false;
   END_IF;
END_FUNCTION_BLOCK

